VERSION : 1.4
// Der FC 53 kann fuer Motoren mit Umrichter, 2 Drehzahlen bzw 2 Punkteverstellung 
// verwendet werden.
// 
// Wird der Baustein mit Umrichter betrieben, so ist das Netzschuetz fuer den 
// Umrichter ans Netz verwendet.
// 
// Wir der Baustein ohne Umrichter betrieben, so ist das Netzschuetz fuer die  
// kleine Drehzahl verwendet.
// 
// Info: Stoerung Laufzeit Speisepumpe. Die eingestellte Zeit in der die 
// Speisepumpe den Pumpenvordruck aufbauen muss ist abgelaufen.
   VAR_INPUT
      IN_ControlVoltage : Bool;   // Delay switch on frequency unit after emergency stop (protection)
      IN_OperationMode_Valid : Bool;   // A valid operation mode (manual or automatic) is selected
      IN_OPerationMode_Active : Bool;   // Opearation mode is selected and hydraulic is active
      IN_Min_PrePressure : Bool;   // Inputsignal pressurelevel of pre pressure pump reached
      IN_Max_PressureComponent : Bool;   // Inputsignal maximum component pressure after pump exceeded
      IN_MotorprotectionPump : Bool;   // Inputsignal error power supply or motor protection of component pump
      IN_With_FU_Pump : Bool;   // Select control of component pump by frequeny unit
      IN_FLT_FU_Pump : Bool;   // Inputsignal fault of frequeny unit component pump
      IN_MaxLevelTray : Bool;   // Input fault max. filling level tray
      IN_Shot_Start : Bool;   // Foaming is active
      IN_MinPressure : Bool;   // Inputsignal fault min pressure of component pump
      IN_PreAlarmBearing : Bool;
      IN_AlarmBearing : Bool;
      IN_Reset_fault_Fkt : Bool;   // Quit faults inside the function block
      IN_ReleaseExternal : Bool;   // External Signal release of pump-/ frequncy unit
      IN_FaultGroup_1 : Bool;   // Fault message of level 1 is active and was not acknowledged
      IN_SOverSOffSWU_running : Bool;   // Switchover- Switchoff- time switch over unit still running
      IN_High_speed : Bool;   // High speed running
      IN_2point_Adjustment : Bool;   // 2 point adjustment is activ
      IN_Cycle_running : Bool;   // Foaming cycle was started and is active
      IN_Recirc_reduced : Bool;   // Reduced recirculation is selected and active
      IN_Recirc_lowpressure : Bool;   // Lowpressure recirculation is selected and active
      IN_Recirc_highpressure : Bool;   // Highpressure recirculation is selected and active
      IN_Recirc_pausetime : Bool;   // Pausetime during interval function active
      IN_UsedForShot : Bool;   // This component will be used for the next part shot
      IN_Delay_Restart : S5Time;   // Time value restart lock of component pump
      IN_Timer_Restart : Timer;   // Timer restart lock of component pump
      IN_RunDownTime_FeedPump : S5Time;   // Time value run down time feed pump
      IN_Timer_ControlFeedPump : Timer;   // Timer of pressure build up control feed pump
      IN_TimerOffFeedPump : Timer;   // Timer to delay switch off from feeding pump
      IN_Timer_Delay_EnClosedL : Timer;   // Timer delay release flow controller
      IN_TimerInterval : Timer;   // Timer for interval times
   END_VAR
   VAR_OUTPUT
      OUT_2_Point_Adjust : Bool;   // Output 2 point adjustment of pump
      OUT_Dosing_active : Bool;   // Signal dosing of component to ProCan-modul
      OUT_Enableclosedloop : Bool;   // Signal of Flow Index "enableclosedloop" to ProCan-modul
      OUT_Pump_MainsContactor : Bool;   // Output mainscontactor pump/frequency unit; or low speed contactor
      OUT_Release_FU : Bool;   // Output release frequency unit; or high speed contactor
   END_VAR
   VAR_IN_OUT
      IO_QPB_Pumpe : Bool;   // Toggelsignal of quick pressure build up to ProCan modul
      IO_Status : ANY;   // Storage of state component pump - state of program block
      IO_Fault : ANY;
      IO_Config : ANY;
      IO_NewFault : Bool;
      IO_FaultLevel_1 : Bool;
      IO_FaultLevel_2 : Bool;
      IO_FaultLevel_3 : Bool;
   END_VAR
   VAR_TEMP
      Temp_IO_Status : "UDT053_Pump";
      ERROR_CODE : Int;   // Error state of systemfunction "BLKMOV" Blockmove
      AnyPointer1 : ANY;   // Pointer to copy the array "IO_Status" and "Temp_IO_Status"
      AnyPointer2 : ANY;   // Pointer to copy the array "IO_Status" and "Temp_IO_Status"
      AnyPointer3 : ANY;   // Pointer to copy the array "IO_Config"
      ReleaseFentingPump : Bool;   // Flag of release fenting pump
      Feedpump_wo_postrun : Bool;   // Flag activation feed pump without component pump post run
      Temp_IO_Fault : "UDT1853_FLT_MeteringPump";
      Temp_IO_Config : "UDT753_MeteringPump";
      ComponentOFF : Bool;   // Component is switched off or on pause time interval
   END_VAR
BEGIN

REGION Network 1: Saved data integration
   // Änderungen:
   // -------------------------------------------------------------------------------
   // Da nach einem sofortigem Widereinschalten der Pumpen nach einer Störung 
   // "STG_Max_Druck" kann es zu einem beschädigen der Pumpen kommen. 
   // Hier wird hier nun über den Weg der Entlüftungspumpe eine Einschaltverzögerung 
   // vorgenommen.
   // 
   // v.d.Geest     20.09.2005
   // -------------------------------------------------------------------------------
   // Auch wenn die Pumpe nicht mit Speisepumpe betrieben wurde wird das Bit 
   // "#Temp_IO_Status.Anforderung_Speisepumpe" gesetzt. 
   // Dieses Signal wurde direkt mit dem Eingang "#IN_Mit_Speisepumpe" verknüpft.
   // 
   // v.d.Geest     16.07.2005
   // -------------------------------------------------------------------------------
   // Der Ausgang "OUT_hohe_Drehzahl" kann entfallen wenn dieser mit dem Ausgang 
   // "#OUT_Freigabe_an_FU_Pumpe" zusammengelegt wird.
   // Bei einem Pumpenstrang ohne Umrichter wäre dieses nun der Ausgang für die hohe 
   // Drehzahl der Pumpen.
   // 
   // Escher        25.11.2004
   // -------------------------------------------------------------------------------
   // Das Signal "Dosieren_an_PUC" war von der Reglerfreigabe an den 
   // Frequenzumrichter abhängig. Die PUC benötigt dieses Signal aber im Schäumzyklus 
   // auch bei ungeregelten Maschinen. (Änderungen im Netzwerk 7)
   // 
   // Strauß        02.08.2004
   // -------------------------------------------------------------------------------
   // Bei einer Verwendung der Komponentenpumpe mit Speisepumpe trat beim ausschalten 
   // der Betriebsart im Kreislauf die Störung "STG_SpP_Laufzeit" auf.
   // Dieses war der Fall wenn die Nachlaufzeit größer eingegeben war als die 
   // Überwachungszeit des Vordrucks.
   // Dieses wurde unterbunden indem die Speisepumpe bei nicht aktiver Betriebsart 
   // nicht mehr angesteuert wird. 
   // Änderungen im Netzwerk 5 durch einfügen von "#IN_Betriebsart_Aktiv" bei der 
   // Zuweisung der "#Temp_IO_Status.Anforderung_Speisepumpe".
   // 
   // v.d.Geest     09.09.2003
   // -------------------------------------------------------------------------------
   // Wenn die Komponentenpumpe ohne Umrichter betrieben wird ist es nicht nötig das 
   // die Anlaufverzögerung nach Steuerspannung Aus abläuft.
   // Deshalb wird das Bit "FRG_UR_wieder_ans_Netz" auch gesetzt, wenn kein Umrichter 
   // verwendet wird. Hierdurch brauch auch die Freigabe für den Zyklus nicht 
   // verändert werden.
   // 
   // v.d.Geest     15.04.2003
   // -------------------------------------------------------------------------------
   // Wenn mehrere Komponentenpumpen mit Speise- oder Entlüftungspumpen betrieben 
   // werden konnte ein unterschiedliches Anlaufen der Komponentenpumpen nur 
   // "außerhalb" des Bausteins unterbunden werden.
   // Hierfür wurde der neue Übergabeparameter "IN_Freigabe_extern" eingebunden. Also 
   // bitte bei einspielen des Bausteins auf die Änderung bim FB achten.
   // 
   // v.d.Geest     11.04.2003
   // -------------------------------------------------------------------------------
   // Um bei größeren Komponentenpumpen auch beim Ausschalten des Kreislaufes oder 
   // nach dem Zyklus ein nichtabreißen des Komponentenstromes zu gewährleisten muß 
   // hier die Speisepumpe, falls vorhanden, nachlaufen.
   // Diese Nachlaufzeit wird von außen vorgegeben sollte aber "fest" bleiben.
   // 
   // Jäger         01.04.2003
   // -------------------------------------------------------------------------------
   // Bei unterschreiten des Min. Füllstandes während des Zyklusses wurde die 
   // Ansteuerung der Materialpumpen abgebrochen.
   // Nur noch ein Abbruch wenn der Zyklus nicht mehr läuft
   // 
   // v.d.Geest     25.02.2003
   // -------------------------------------------------------------------------------
   // Die Störung des Vordruckes wird unabhängig von der Anforderung ausgewertet.
   // Hierdurch wird ein kurzes Anlaufen der Materialpumpnen bei nicht vorhandenen 
   // Vordruck unterbunden.
   // 
   // Lindner       27.01.2003
   // -------------------------------------------------------------------------------
         LAR1;
         L;
         LAR2;
   //
         L     W[AR2, P#0.0];  // Bytes
         T     W[AR1, P#0.0];
         L     W[AR2, P#2.0];  //Amount of bytes
         T     W[AR1, P#2.0];
         L     W[AR2, P#4.0];  //Block no,
         T     W[AR1, P#4.0];
         L     D[AR2, P#6.0];  //Startadress of datas
         T     D[AR1, P#6.0];
   //
         CALL  BLKMOV
         ( SRCBLK  := #AnyPointer1,
           RET_VAL := #ERROR_CODE,
           DSTBLK  := #Temp_IO_Status
         );
   //
         LAR1;
         L;
         LAR2;
   //
         L     W[AR2, P#0.0];  // Bytes
         T     W[AR1, P#0.0];
         L     W[AR2, P#2.0];  //Amount of bytes
         T     W[AR1, P#2.0];
         L     W[AR2, P#4.0];  //Block no,
         T     W[AR1, P#4.0];
         L     D[AR2, P#6.0];  //Startadress of datas
         T     D[AR1, P#6.0];
   //
         CALL  BLKMOV
         ( SRCBLK  := #AnyPointer2,
           RET_VAL := #ERROR_CODE,
           DSTBLK  := #Temp_IO_Fault
         );
   //
   //
         LAR1;
         L;
         LAR2;
   //
         L     W[AR2, P#0.0];  // Bytes
         T     W[AR1, P#0.0];
         L     W[AR2, P#2.0];  //Amount of bytes
         T     W[AR1, P#2.0];
         L     W[AR2, P#4.0];  //Block no,
         T     W[AR1, P#4.0];
         L     D[AR2, P#6.0];  //Startadress of datas
         T     D[AR1, P#6.0];
   //
         CALL  BLKMOV
         ( SRCBLK  := #AnyPointer3,
           RET_VAL := #ERROR_CODE,
           DSTBLK  := #Temp_IO_Config
         );
END_REGION

REGION Network 2: Handle interval mode
   // Messages
         A     #Temp_IO_Config.PumpDeselectedInterval;
         FP    #Temp_IO_Status.Mes_PumpDeselectedInt;
         R     #Temp_IO_Config.PumpDeselected;
         A     #Temp_IO_Config.PumpDeselected;
         FP    #Temp_IO_Status.Mes_PumpDeselected;
         R     #Temp_IO_Config.PumpDeselectedInterval;

         A     #Temp_IO_Status.Mes_PumpDeselectedInt;
         =     #Temp_IO_Fault.Mes_PumpDeselectedInt;
         A     #Temp_IO_Status.Mes_PumpDeselected;
         =     #Temp_IO_Fault.Mes_PumpDeselected;

         AN    #Temp_IO_Config.PumpDeselectedInterval;
         R     #Temp_IO_Status.IntervalPause;

   // Interval times
         A     #Temp_IO_Config.PumpDeselectedInterval;
         FP    #Temp_IO_Status.HF_FPPumpDeselectedInt;
         JCN   int;
         R     #Temp_IO_Status.IntervalPause;
         CLR;
         L     S5T#0MS;
         SP    #IN_TimerInterval;
         JU    eint;

   int:  AN    #Temp_IO_Config.PumpDeselectedInterval;
         JC    eint;

   // Change run time <-> pause time
         AN    #IN_TimerInterval;
         JCN   eint;

   // Select the correct time
         L     #Temp_IO_Config.RunTimePumpInterval;
         A     #Temp_IO_Status.IntervalPause;
         JC    time;
         L     #Temp_IO_Config.PauseTimePumpInterval;

   // Start timer
   time: CLR;
         SE    #IN_TimerInterval;
         SET;
         SE    #IN_TimerInterval;
         AN    #Temp_IO_Status.IntervalPause;
         =     #Temp_IO_Status.IntervalPause;
   eint: NOP   0;
   // switch off if necessary
         O     #Temp_IO_Config.PumpDeselected;
         O     #Temp_IO_Status.IntervalPause;
         =     #ComponentOFF;
END_REGION

REGION Network 3: Switch on delay of frequency unit
   // Bei Betrieb mit Umrichter wird der Umrichter mit einer Wiedereinschaltsperre 
   // von 30 Sek. geschützt. Nach Steuerspannung AUS wird der Umrichter 30 Sek. lang 
   // vom Netz getrennt auch wenn die Steuerspannung sofort wieder eingeschaltet 
   // wird.
   //--------- Frequency unit back to power supply ---------------
   //      O     #Temp_IO_Status.FLT_Max_pressure    // Bitte testen 25.6.08 HK
         AN    #IN_ControlVoltage;
         AN    #ComponentOFF;
         O     #ComponentOFF;
         FP    #Temp_IO_Status.Rampe_Voltage_Off;
         R     #Temp_IO_Status.Release_Startup_FC;
         R     #IN_Timer_Restart;
         R     #Temp_IO_Status.Start_Startupdelay;
   //
         A     #Temp_IO_Status.Release_Startup_FC;
         JC    Run;
   //
         A     #Temp_IO_Status.Start_Startupdelay;
         AN    #Temp_IO_Status.Release_Startup_FC;
         L     S5T#10S;
         SD    #IN_Timer_Restart;
   //
         SET;
         S     #Temp_IO_Status.Start_Startupdelay;
   //
         O     #IN_Timer_Restart;
         ON    #IN_With_FU_Pump;
         S     #Temp_IO_Status.Release_Startup_FC;
         R     #IN_Timer_Restart;
         R     #Temp_IO_Status.Start_Startupdelay;
   //
   Run:  NOP   0;
END_REGION

REGION Network 4: Fault handling
   //--------- Störung Reset --------------------------
         A     #IN_Reset_fault_Fkt;
         R     #Temp_IO_Fault.FLT_Prepressure;
         R     #Temp_IO_Fault.FLT_Motorprotection;
         R     #Temp_IO_Fault.FLT_Max_pressure;
         R     #Temp_IO_Fault.FLT_SpP_Runtime;
         R     #Temp_IO_Fault.FLT_F_converter;
         R     #Temp_IO_Fault.FLT_Min_Pressure;
         R     #Temp_IO_Fault.FLT_DeselectedCompReqest;
         R     #Temp_IO_Fault.FLT_MaxLTripTray;
         R     #Temp_IO_Fault.FLT_PreAlarmBearing;
         R     #Temp_IO_Fault.FLT_AlarmBearing;
   //--------- Störung Pumpenvordruck -----------------
         A     #Temp_IO_Status.Netrelais;
         AN    #IN_Min_PrePressure;
         AN    #IN_With_FU_Pump;
         O;
         A     #IN_With_FU_Pump;
         A     #Temp_IO_Status.Controllrelease_to_FC;
         AN    #IN_Min_PrePressure;
         O;
         AN    #Temp_IO_Config.WithFeedPump;
         AN    #IN_Min_PrePressure;
         AN    #ComponentOFF;
         AN    #Temp_IO_Fault.FLT_Prepressure;
         S     #Temp_IO_Fault.FLT_Prepressure;
         S     #IO_NewFault;
   //--------- Störung Laufzeit Speisepumpe -----------
         A     #Temp_IO_Status.Selection_Feedingpump;
         A     #Temp_IO_Config.WithFeedPump;
         AN    #IN_Min_PrePressure;
         L     #Temp_IO_Config.DelayPressureFeedP;
         SD    #IN_Timer_ControlFeedPump;
   //
         A     #IN_Timer_ControlFeedPump;
         AN    #Temp_IO_Fault.FLT_SpP_Runtime;
         S     #Temp_IO_Fault.FLT_SpP_Runtime;
         S     #IO_NewFault;
   //--------- Störung Motorschutz --------------------
         A     #IN_MotorprotectionPump;
         AN    #ComponentOFF;
         AN    #Temp_IO_Fault.FLT_Motorprotection;
         S     #Temp_IO_Fault.FLT_Motorprotection;
         S     #IO_NewFault;
   //--------- Störung max. Druck  --------------------
         AN    #IN_Max_PressureComponent;
         AN    #ComponentOFF;
         AN    #Temp_IO_Fault.FLT_Max_pressure;
         S     #Temp_IO_Fault.FLT_Max_pressure;
         S     #IO_NewFault;
   //--------- Fault deselected component requested for shot  ---
         O     #Temp_IO_Config.PumpDeselectedInterval;
         O     #Temp_IO_Config.PumpDeselected;
         A     #IN_UsedForShot;
         AN    #Temp_IO_Fault.FLT_DeselectedCompReqest;
         S     #Temp_IO_Fault.FLT_DeselectedCompReqest;
         S     #IO_NewFault;
   //--------- Störung Umrichter  ---------------------
         ON    #IN_With_FU_Pump;
         ON    #Temp_IO_Status.Release_Startup_FC;
         O     #ComponentOFF;
         JC    K_UR;
         A     #Temp_IO_Status.Netrelais;
         L     S5T#15S;
         SD    #IN_Timer_Restart;
         A     #IN_Timer_Restart;
         AN    #IN_FLT_FU_Pump;
         AN    #Temp_IO_Fault.FLT_F_converter;
         S     #Temp_IO_Fault.FLT_F_converter;
         S     #IO_NewFault;

   //-----
         AN    #IN_MaxLevelTray;
         AN    #Temp_IO_Fault.FLT_MaxLTripTray;
         S     #Temp_IO_Fault.FLT_MaxLTripTray;
         S     #IO_NewFault;

   K_UR: NOP   0;
   //--------- Min pressure at     -------------------
   //---------  shot start         -------------------
         A     #IN_Shot_Start;
         AN    #IN_MinPressure;
         A     #IN_UsedForShot;
         AN    #Temp_IO_Fault.FLT_Min_Pressure;
         S     #Temp_IO_Fault.FLT_Min_Pressure;
         S     #IO_NewFault;

         A     #IN_PreAlarmBearing;
         AN    #Temp_IO_Fault.FLT_PreAlarmBearing;
         S     #Temp_IO_Fault.FLT_PreAlarmBearing;
         S     #IO_NewFault;

         A     #IN_AlarmBearing;
         AN    #Temp_IO_Fault.FLT_AlarmBearing;
         S     #Temp_IO_Fault.FLT_AlarmBearing;
         S     #IO_NewFault;

         A     #Temp_IO_Status.Start_Startupdelay;
         =     #Temp_IO_Fault.Mes_StartUpDelayFU;
END_REGION

REGION Network 5: Error handling fault groups
         O     #Temp_IO_Fault.FLT_Prepressure;
         O     #Temp_IO_Fault.FLT_Motorprotection;
         O     #Temp_IO_Fault.FLT_Max_pressure;
         O     #Temp_IO_Fault.FLT_F_converter;
         O     #Temp_IO_Fault.FLT_SpP_Runtime;
         O     #Temp_IO_Fault.FLT_Min_Pressure;
         O     #Temp_IO_Fault.FLT_DeselectedCompReqest;
         O     #Temp_IO_Fault.FLT_AlarmBearing;
         O     #Temp_IO_Fault.FLT_MaxLTripTray;
         S     #IO_FaultLevel_1;

   //      O     XXXXXXXX
   //      S     #IO_FaultLevel_2

         O     #Temp_IO_Fault.FLT_PreAlarmBearing;
         S     #IO_FaultLevel_3;
   //
         O     #Temp_IO_Fault.FLT_Prepressure;
         O     #Temp_IO_Fault.FLT_Motorprotection;
         O     #Temp_IO_Fault.FLT_Max_pressure;
         O     #Temp_IO_Fault.FLT_F_converter;
         O     #Temp_IO_Fault.FLT_SpP_Runtime;
         O     #Temp_IO_Fault.FLT_Min_Pressure;
         O     #Temp_IO_Fault.FLT_DeselectedCompReqest;
         O     #Temp_IO_Fault.FLT_AlarmBearing;
         O     #Temp_IO_Fault.FLT_PreAlarmBearing;
         O     #Temp_IO_Fault.FLT_MotorFan;
         O     #Temp_IO_Fault.FLT_MaxLTripTray;
         =     #Temp_IO_Status.FLT_Exist;
END_REGION

REGION Network 6: Venting pump
   //       ON    #Temp_IO_Status.STG_Min_Level
   //       O     #IN_Cycle_running
   //     U     #IN_Mit_Entlueftungspumpe
   //       U     #IN_OperationMode_Valid
   //       UN    #Temp_IO_Fault.FLT_Prepressure
   //       =     #Freigabe_Enlt_Pumpe
   //
   //      U     #Temp_IO_Status.Ventingtime_finished
   //      SPB   P_ok
   //
   //      U     #Freigabe_Enlt_Pumpe
   //      L     S5T#10S
   //      SE    #IN_Timer_Universal
   //-------------------------------------------------
   //       O     #IN_Timer_Universal
   //       ON    #IN_Mit_Entlueftungspumpe
   //       S     #Temp_IO_Status.Ventingtime_finished
   //-------------------------------------------------
   //      SPBN  P_ok
   //
   //       CLR
   //       SI    #IN_Timer_Universal
   //
   // P_ok: NOP 0
   //-------------------------------------------------
   //       U     #Temp_IO_Status.STG_Min_Level
   //       UN    #IN_Cycle_running
   //       ON    #IN_ControlVoltage
   //       O     #Temp_IO_Fault.FLT_Prepressure
   //       R     #Temp_IO_Status.Ventingtime_finished
   //-------------------------------------------------
   //      ON    #Temp_IO_Status.Ventingtime_finished
   //       O     #Temp_IO_Status.Allg_Pumpenanforderung
   //       U     #Freigabe_Enlt_Pumpe
   //       UN    #Temp_IO_Status.STG_Motorsch_Entl_Pumpe
   //       =     #Temp_IO_Status.Netzschuetz_Entl_Pumpe
END_REGION

REGION Network 7: Pump
         O     #IN_Recirc_reduced;
         O     #IN_Recirc_lowpressure;
         A(;
         ON    #IN_Recirc_pausetime;
         O     #IN_Cycle_running;
         );
         O     #IN_Recirc_highpressure;
         O     #IN_Cycle_running;
         A     #IN_OPerationMode_Active;
         AN    #IN_FaultGroup_1;
         AN    #Temp_IO_Fault.FLT_Prepressure;
         AN    #Temp_IO_Fault.FLT_Motorprotection;
         AN    #Temp_IO_Fault.FLT_Max_pressure;
         AN    #Temp_IO_Fault.FLT_SpP_Runtime;
         AN    #Temp_IO_Fault.FLT_F_converter;
   //      U     #Temp_IO_Status.Ventingtime_finished
         A     #IN_ControlVoltage;
         AN    #ComponentOFF;
         =     #Feedpump_wo_postrun;
         A     #Feedpump_wo_postrun;
         L     #IN_RunDownTime_FeedPump;
         SF    #IN_TimerOffFeedPump;
   //
         A     #IN_TimerOffFeedPump;
         A     #Temp_IO_Config.WithFeedPump;
         A     #IN_OPerationMode_Active;
         =     #Temp_IO_Status.Selection_Feedingpump;
   //-------------------------------------------------
         ON    #Temp_IO_Status.Release_Startup_FC;
         O     #IN_With_FU_Pump;
         JC    Allg;
         AN    #IN_With_FU_Pump;
         A     #Temp_IO_Status.High_rpm;
         AN    #IN_High_speed;
         L     #IN_Delay_Restart;
         SE    #IN_Timer_Restart;
   //-------------------------------------------------
   Allg: AN    #IN_With_FU_Pump;
         A     #Feedpump_wo_postrun;
         A     #IN_Min_PrePressure;
         AN    #IN_Timer_Restart;
         O;
         A     #IN_With_FU_Pump;
         A     #Feedpump_wo_postrun;
         A     #IN_Min_PrePressure;
         =     #Temp_IO_Status.Main_Pumpselection;
   //------ Umrichter ans Netz bzw. kleine Drehzahl --
         A     #IN_ReleaseExternal;
         A     #Temp_IO_Status.Main_Pumpselection;
         AN    #IN_With_FU_Pump;
         O;
         A     #IN_With_FU_Pump;
         A     #IN_ControlVoltage;
         AN    #ComponentOFF;
         A     #Temp_IO_Status.Release_Startup_FC;
         =     #Temp_IO_Status.Netrelais;
   //-------------------------------------------------
         O     #IN_Recirc_reduced;
         O     #IN_Recirc_lowpressure;
         A(;
         ON    #IN_Recirc_pausetime;
         O     #IN_Cycle_running;
         );
         O     #IN_Recirc_highpressure;
         O     #IN_Cycle_running;
         A     #IN_ReleaseExternal;
         A     #Temp_IO_Status.Main_Pumpselection;
         AN    #Temp_IO_Fault.FLT_Prepressure;
         AN    #Temp_IO_Fault.FLT_Motorprotection;
         AN    #Temp_IO_Fault.FLT_Max_pressure;
         AN    #Temp_IO_Fault.FLT_SpP_Runtime;
         AN    #Temp_IO_Fault.FLT_F_converter;
         A     #IN_FLT_FU_Pump;
         =     #Temp_IO_Status.Controllrelease_to_FC;
END_REGION

REGION Network 8: High speed and 2 point adjustment if drive without FU
         A     #Temp_IO_Status.Netrelais;
         A     #IN_High_speed;
         =     #Temp_IO_Status.High_rpm;
   //-------------------------------------------------
         A     #Feedpump_wo_postrun;
         A     #IN_2point_Adjustment;
         =     #Temp_IO_Status.Valve_2_point_selection;
END_REGION

REGION Network 9: Release of controller to modul of machine
         A     #IN_ReleaseExternal;
         A     #Temp_IO_Status.Main_Pumpselection;
         AN    #IN_With_FU_Pump;
         O     #Temp_IO_Status.Controllrelease_to_FC;
         =     #Temp_IO_Status.Metering_to_PUC;
   //
         A     #Temp_IO_Status.Controllrelease_to_FC;
         L     S5T#300MS;
         SD    #IN_Timer_Delay_EnClosedL;

         A     #IN_Timer_Delay_EnClosedL;
         =     #Temp_IO_Status.Enableclosedloop;
END_REGION

REGION Network 10: Quick pressure build up
   // Nur notwendig fuer "Schnellen Druckaufbau" mit Modul !!!
         O     #IN_Cycle_running;
         O     #IN_Recirc_highpressure;
         A     #IN_With_FU_Pump;
         AN    #IN_SOverSOffSWU_running;
         A     #Temp_IO_Status.Enableclosedloop;
         A(;
         O     #IN_UsedForShot;
         ON    #IN_Cycle_running;
         );
         FP    #Temp_IO_Status.Puls_SDA;
         JCN   SDA;
         AN    #IO_QPB_Pumpe;
         =     #IO_QPB_Pumpe;
   SDA:  NOP   0;
END_REGION

REGION Network 11: Allocation of outputs
         A     #Temp_IO_Status.Netrelais;
         =     #OUT_Pump_MainsContactor;
   //-------------------------------------------------
         A     #Temp_IO_Status.Valve_2_point_selection;
         =     #OUT_2_Point_Adjust;
   //-------------------------------------------------
         A     #Temp_IO_Status.Controllrelease_to_FC;
         A     #IN_With_FU_Pump;
         O;
         A     #Temp_IO_Status.High_rpm;
         AN    #IN_With_FU_Pump;
         =     #OUT_Release_FU;
   //-------------------------------------------------
         A     #Temp_IO_Status.Metering_to_PUC;
         =     #OUT_Dosing_active;
   //-------------------------------------------------
         A     #IN_With_FU_Pump;
         A     #Temp_IO_Status.Enableclosedloop;
         =     #OUT_Enableclosedloop;
   //-------------------------------------------------
END_REGION

REGION Network 12: Function is active
         SET;
         =     #Temp_IO_Status.Block_is_active;
END_REGION

REGION Network 13: Save data
         CALL  BLKMOV
         ( SRCBLK  := #Temp_IO_Status,
           RET_VAL := #ERROR_CODE,
           DSTBLK  := #AnyPointer1
         );
   //
         CALL  BLKMOV
         ( SRCBLK  := #Temp_IO_Fault,
           RET_VAL := #ERROR_CODE,
           DSTBLK  := #AnyPointer2
         );
   //
         CALL  BLKMOV
         ( SRCBLK  := #Temp_IO_Config,
           RET_VAL := #ERROR_CODE,
           DSTBLK  := #AnyPointer3
         );
END_REGION
END_FUNCTION

FUNCTION "FC054_FaultsMetering" : Void   // FC54, STL
TITLE = Faults ProCan flowstate
{ S7_Optimized_Access := 'FALSE' }
NAME : Fault
VERSION : 0.1
   VAR_INPUT
      IN_ProCanFlow_State : Struct
         Flowstopped : Bool;   // piston has stopped
         FlowQPB : Bool;   // Flow quick pressure build up is active
         ControlOnUpperLimit : Bool;   // flow control loop operates on it upper limits
         ControlOnLowerLimit : Bool;   // flow control loop operates on its lower limits
         FlowtoleranceL : Bool;   // tolerance: flow is too low
         FlowtoleranceH : Bool;   // tolerance: flow is too high
      END_STRUCT;
      IN_Reset_Fault : Bool;
   END_VAR
   VAR_IN_OUT
      IO_Any_Flow_Fault : ANY;
      IO_HF_FLT_QPB : Bool;
      IO_FaultLevel1 : Bool;
      IO_FaultLevel2 : Bool;
      IO_FaultLevel3 : Bool;
      IO_NewFault : Bool;
   END_VAR
   VAR_TEMP
      Temp_Any_Flow_Fault : ANY;
      Temp_Flow_Fault : "UDT1853_FLT_MeteringPump";
      ERROR_CODE : Int;
      Temp_FLT_Tolerance_high : Bool;
      Temp_FLT_Tolerance_low : Bool;
      Temp_FLT_FlowContrAtLim : Bool;
      Temp_Flt_FlowSDAtimeOut : Bool;
   END_VAR
BEGIN

REGION Network 1: Get temporary variables flow fault
         L;
         LAR1;
         LAR2;
   //
         L     W[AR1, P#0.0];  // Bytes
         T     W[AR2, P#0.0];
         L     W[AR1, P#2.0];  // Amount of bytes
         T     W[AR2, P#2.0];
         L     W[AR1, P#4.0];  // Block no,
         T     W[AR2, P#4.0];
         L     D[AR1, P#6.0];  // Startadress of data
         T     D[AR2, P#6.0];
   //
         CALL  BLKMOV
         ( SRCBLK  := #Temp_Any_Flow_Fault,
           RET_VAL := #ERROR_CODE,
           DSTBLK  := #Temp_Flow_Fault
         );
END_REGION

REGION Network 2: Reset faults flow
         AN    #IN_Reset_Fault;
         JC    nw3e;

         CLR;
         =     #Temp_Flow_Fault.FLT_Tolerance_high;
         =     #Temp_Flow_Fault.FLT_Tolerance_low;
         =     #Temp_Flow_Fault.FLT_FlowControlAtLimit;
         =     #Temp_Flow_Fault.FLT_FlowControlAtLOWLimit;
         =     #Temp_Flow_Fault.FLT_FlowSDATimeOut;

   nw3e: NOP   0;
END_REGION

REGION Network 3: Fault flow state of ProCan module
   //      L     #IN_ProCanFlow_State
   //      L     16
   //      UW
   //      L     0
   //      <>D
   //      FP    #IO_HF_FLT_QPB
   //      =     #Temp_Flt_FlowSDAtimeOut

   //      U     #Temp_Flt_FlowSDAtimeOut
   //      UN    #Temp_Flow_Fault.FLT_FlowSDATimeOut
   //      S     #Temp_Flow_Fault.FLT_FlowSDATimeOut
   //      S     #IO_NewFault

         A     #IN_ProCanFlow_State.ControlOnUpperLimit;
         AN    #Temp_Flow_Fault.FLT_FlowControlAtLimit;
         S     #Temp_Flow_Fault.FLT_FlowControlAtLimit;
         S     #IO_NewFault;

         A     #IN_ProCanFlow_State.ControlOnLowerLimit;
         AN    #Temp_Flow_Fault.FLT_FlowControlAtLOWLimit;
         S     #Temp_Flow_Fault.FLT_FlowControlAtLOWLimit;
         S     #IO_NewFault;
END_REGION

REGION Network 4: Fault levels
   //    O     xxxxxxxxx
   //    =     #IO_FaultLevel1

         O     #Temp_Flow_Fault.FLT_Tolerance_high;
         O     #Temp_Flow_Fault.FLT_Tolerance_low;
         O     #Temp_Flow_Fault.FLT_FlowControlAtLimit;
         O     #Temp_Flow_Fault.FLT_FlowControlAtLOWLimit;
         O     #Temp_Flow_Fault.FLT_FlowSDATimeOut;
         S     #IO_FaultLevel3;
END_REGION

REGION Network 5: Write back faults
         CALL  BLKMOV
         ( SRCBLK  := #Temp_Flow_Fault,
           RET_VAL := #ERROR_CODE,
           DSTBLK  := #Temp_Any_Flow_Fault
         );
END_REGION
END_FUNCTION

FUNCTION "FC055_PumpVentilation" : Void   // FC55, STL
TITLE = Function for organize pump Ventilation
{ S7_Optimized_Access := 'FALSE' }
VERSION : 0.1
   VAR_INPUT
      IN_Reset_fault_Fkt : Bool;   // Quit faults inside the function block
      IN_Motorprotection : Bool;   // Inputsignal error power supply or motor protection
      IN_ComponentDeselected : Bool;   // Is the component deselected? -> Fault Group 2 -> Groupe 3
      In_Start : Bool;   // Start value for the ventilation
      IN_Time : S5Time;   // Time value delay switch off the ventilation
      IN_Timer : Timer;   // Timer for delay time to switch off the ventilation
   END_VAR
   VAR_OUTPUT
      OUT_MainContactor : Bool;   // Output maincontactor Ventilation
   END_VAR
   VAR_IN_OUT
      IO_FLT_MotorFan : Bool;
      IO_NewFault : Bool;
      IO_FaultLevel_2 : Bool;
      IO_FaultLevel_3 : Bool;
   END_VAR
BEGIN

REGION Network 1: Fault handling
   //--------- Reset fault ---------------------------
         A     #IN_Reset_fault_Fkt;
         R     #IO_FLT_MotorFan;
   //--------- Fault Motorprotection -----------------
         A     #IN_Motorprotection;
         AN    #IO_FLT_MotorFan;
         S     #IO_FLT_MotorFan;
         S     #IO_NewFault;
   //--------- If selected fault group 2 -------------
         A     #IO_FLT_MotorFan;
         AN    #IN_ComponentDeselected;
         S     #IO_FaultLevel_2;
   //--------- If deselected fault group 3 -----------
         A     #IO_FLT_MotorFan;
         A     #IN_ComponentDeselected;
         S     #IO_FaultLevel_3;
   //-------------------------------------------------
END_REGION

REGION Network 2: Start venting
   //-----
         A     #In_Start;
         AN    #IO_FLT_MotorFan;
         L     #IN_Time;
         SF    #IN_Timer;
         A     #IN_Timer;
         AN    #IO_FLT_MotorFan;
         =     #OUT_MainContactor;
   //-----
END_REGION
END_FUNCTION

FUNCTION "FC056_TemPulse2" : Void   // FC56, STL
TITLE = Temperature control pulse width
{ S7_Optimized_Access := 'FALSE' }
VERSION : 0.1
   VAR_INPUT
      Trig : Bool;
      In_Sollwert : Real;
      In_Istwert_Tank : Real;
      In_Istwert_Return : Real;
      In_Wichtung : Real;
      In_Regelstrecke : Real;
      In_MaxDelta_K : Real;
      In_MaxDelta_H : Real;
   END_VAR
   VAR_IN_OUT
      Pulsezeit : Real;
      Heating : Bool;
      Cooling : Bool;
   END_VAR
   VAR_TEMP
      Value1 : Real;
      Value2 : Real;
      Value3 : Real;
      Value4 : Real;
      Value5 : Real;
      Value6 : Real;
      Value7 : Real;
      MaxDelta : Real;
      Istwert_Tank : Real;
      Istwert_Return : Real;
      Sollwert : Real;
      Wichtung : Real;
      MaxDelta_K : Real;
      MaxDelta_H : Real;
      Regelstrecke : Real;
      Pulsezeit_real : Real;
   END_VAR
BEGIN

REGION Network 1: Berechnen nur wenn Timer abgelaufen
         AN    #Trig;
         BEC;
END_REGION

REGION Network 2: Werte wandeln von INT in REAL
         L     #In_Sollwert;
         T     #Sollwert;

         L     #In_Istwert_Tank;
         T     #Istwert_Tank;

         L     #In_Istwert_Return;
         T     #Istwert_Return;

         L     #In_Wichtung;
         T     #Wichtung;

         L     #In_Regelstrecke;
         T     #Regelstrecke;

         L     #In_MaxDelta_K;
         T     #MaxDelta_K;

         L     #In_MaxDelta_H;
         T     #MaxDelta_H;
END_REGION

REGION Network 3: Mittelwert bilden
         L     #Istwert_Tank;
         L     #Wichtung;
         *R;
         T     #Value1;

         L     100.0;
         L     #Wichtung;
         -R;
         L     #Istwert_Return;
         *R;
         T     #Value2;

         L     #Value1;
         L     #Value2;
         +R;
         L     100.0;
         /R;
         T     #Value3;  // Mittelwert
END_REGION

REGION Network 4
   // Ist dieser Wert negativ, dann mit MaxDelta_H arbeiten
         L     #Value3;
         L     #Sollwert;
         -R;
         T     #Value4;  // Differenz Mittelist - Sollwert

         L     #MaxDelta_K;  // Wert für Kühlen
         T     #MaxDelta;

         L     #Value4;
         L     0;
         <R;
         JCN   Limi;
         L     #MaxDelta_H;  // Für Heizen diesen Wert nehmen
         T     #MaxDelta;
END_REGION

REGION Network 5
   // Differenz auf MaxWert limitieren
   Limi: L     #Value4;
         L     #MaxDelta;
         >R;
         JCN   kMax;
         T     #Value5;
         JU    calc;

   kMax: L     #Value4;
         T     #Value5;
END_REGION

REGION Network 6
   calc: NOP   0;

         L     100.0;
         L     #Value5;
         *R;
         L     #MaxDelta;
         /R;
         T     #Value6;
END_REGION

REGION Network 7: Pulsezeit: - >> HEIZEN / + >> KÜHLEN
         L     #Regelstrecke;
         L     100.0;
         /R;
         L     #Value6;
         *R;
         T     #Value7;

         L     #Value7;
         L     100.0;
         *R;
         T     #Pulsezeit_real;

   // Wenn noch nicht Positiv, dann machen !
         L     #Pulsezeit_real;
         L     0.0;
         <R;
         JCN   tak;
         L     #Pulsezeit_real;
         NEGR;
         JU    rnd;

   tak:  TAK;
   rnd:  NOP   0;
         L     10.0;
         *R;
         T     #Pulsezeit;  // Ausgabe int INT, aber gleich positiv!
END_REGION

REGION Network 8: Steuerbits ausgeben
         L     #Pulsezeit_real;
         L     0.0;
         >R;
         =     #Cooling;

         L     #Pulsezeit_real;
         L     0.0;
         <R;
         =     #Heating;
END_REGION
END_FUNCTION

FUNCTION "FC057_HPHeatexchanger" : Void   // FC57, STL
{ S7_Optimized_Access := 'FALSE' }
VERSION : 0.1
   VAR_TEMP
      DINT_dummy : Real;
      Imp_WT_Aus : Bool;
      Imp_WT_Ein : Bool;
      Temp_Cooling : Bool;
      Dummy : Bool;
      Temp_MoreDelta : Bool;
      Temp_HD_WT : Real;
      Temp_SetValueTemp : Real;
      Regelstrecke : Time;
      Zeit_abgelaufen : Time;
   END_VAR
BEGIN

REGION Network 1: There is no connection to the sensor (3)
   //---------------------------------------------
   //  Controller temperature Heatexchanger K1
   //---------------------------------------------
         AN    "DB753_MeteringPump".Pump[1].WithHPHeatExchanger;
         R     "DB823_Error_Metering".Temperature_HeatexchangerHP[1].Sensor_FLT_broken_wire;
         R     "DB823_Error_Metering".Temperature_HeatexchangerHP[1].Warning_limit_plus;
         R     "DB823_Error_Metering".Temperature_HeatexchangerHP[1].Warning_limit_minus;
         R     "DB823_Error_Metering".Temperature_HeatexchangerHP[1].Alarm_limit_plus;
         R     "DB823_Error_Metering".Temperature_HeatexchangerHP[1].Alarm_limit_minus;
         R     "DB613_Komponent_State".HeatexchangerHP[1].Fault_Exist;
         JC    EHD1;
   //-----
         CALL  "FC920_PV_Calc_Act_Value"
         ( IN_Act_Value_read := TRUE,
           IN_Act_Value_ext  := FALSE,
           IN_Ext_Value      := #DINT_dummy,
           IN_Read_Double    := FALSE,
           IN_FLT_Needful    := 1,
           IN_FLT_Reset      := "DB009_Faults".Faults_Reset_FKT_M1,
           IO_Any_ArrayPV    := "DB608_PV_Metering".HeatexchangerHP[1],
           IO_Fault_Sensor   := "DB823_Error_Metering".Temperature_HeatexchangerHP[1].Sensor_FLT_broken_wire,
           IO_New_Fault      := "DB009_Faults".Faultschanging_M1,
           IO_FLT_Level_3    := "DB009_Faults".Faults_FKT_Grp_3_M1
         );

   //---------------------------------------------
   //  Controller temperature Heatexchanger K1
   //---------------------------------------------
         L     "DB608_PV_Metering".HeatexchangerHP[1].PV_ActV.Value;
         L     10.0;
         /R;
         T     #Temp_HD_WT;
   //
         L     "DB608_PV_Metering".HeatexchangerHP[1].PV_SetV.Value;
         L     10.0;
         /R;
         T     #Temp_SetValueTemp;
   //
         CALL  "FC056_TemPulse2"
         ( Trig              := "Start_Controler1_HP_K1",
           In_Sollwert       := #Temp_SetValueTemp,
           In_Istwert_Tank   := #Temp_HD_WT,
           In_Istwert_Return := #Temp_HD_WT,
           In_Wichtung       := "DB751_auxiliaryDriveMetering".HeatexchangerHP[1].Weighting_Temp,
           In_Regelstrecke   := "DB751_auxiliaryDriveMetering".HeatexchangerHP[1].PLC_Control_Area,
           In_MaxDelta_K     := "DB751_auxiliaryDriveMetering".HeatexchangerHP[1].Max_Temp_Diff_Cooling,
           In_MaxDelta_H     := "DB751_auxiliaryDriveMetering".HeatexchangerHP[1].Max_Temp_Diff_Heating,
           Pulsezeit         := "DB613_Komponent_State".HeatexchangerHP[1].PulsTime,
           Heating           := #Dummy,
           Cooling           := #Temp_Cooling
         );
   //
   //Regelstrecke ms Format
         L     "DB751_auxiliaryDriveMetering".HeatexchangerHP[1].PLC_Control_Area;
         L     1000.0;
         *R;
         RND;
         T     #Regelstrecke;  // Zeitwert für Timer

   // Regelstreckentimer ständig starten

         AN    "Start_Controler1_HP_K1";
         =     "Start_Controler2_HP_K1";

         CALL  TON , "DB55_Temp_HD_WT_MK1_K1"
         ( IN := "Start_Controler2_HP_K1",
           PT := #Regelstrecke,
           Q  := "Start_Controler1_HP_K1",
           ET := #Zeit_abgelaufen
         );

   // Kühlen  EIN
         A     #Temp_Cooling;
         S     "DB613_Komponent_State".HeatexchangerHP[1].CoolingActive;

   // Kleine Einschatverzögerung
         L     #Temp_SetValueTemp;
         L     "DB751_auxiliaryDriveMetering".HeatexchangerHP[1].Offset_Cooling;
         +R;
         L     #Temp_HD_WT;
         >R;
         =     #Temp_MoreDelta;
   // Kühlen  AUS
         L     "DB613_Komponent_State".HeatexchangerHP[1].PulsTime;
         RND;
         L     #Zeit_abgelaufen;
         <D;
         AN(;
         L     "DB613_Komponent_State".HeatexchangerHP[1].PulsTime;
         RND;
         L     #Regelstrecke;
         >D;
         );
         ON    "DB613_Komponent_State".HeatexchangerHP[1].Switch_Temp_ON_OFF;
         ON    "DB619_State_MPart".Operationmode[1].valid;
         O     "DB823_Error_Metering".Temperature_HeatexchangerHP[1].Sensor_FLT_broken_wire;
         O     #Temp_MoreDelta;
         R     "DB613_Komponent_State".HeatexchangerHP[1].CoolingActive;

         A     "DB613_Komponent_State".HeatexchangerHP[1].CoolingActive;
         A     "DB619_State_MPart".Machine[1].Metering."01";

         =     "V_HP_Heater_Cooling_C1";  // "V_HExchang_Cooling_K1" // stromlos zu
         =     "V_HP_Heater_Bypass_C1";  // "V_HExchang_Bypass_K1" // stromlos offen

   //-----
   // Check limits temperature 1 Heatexchanger

         CALL  "FC916_PV_Limits"
         ( IN_Tolerance_Test     := "DB619_State_MPart".Operationmode[1].Controllvoltage,
           IN_Reset_Fault        := "DB009_Faults".Faults_Reset_FKT_M1,
           IO_Any_ArrayPV        := "DB608_PV_Metering".HeatexchangerHP[1],
           IO_Fault_Warn_upperL  := "DB823_Error_Metering".Temperature_HeatexchangerHP[1].Warning_limit_plus,
           IO_Fault_Warn_lowerL  := "DB823_Error_Metering".Temperature_HeatexchangerHP[1].Warning_limit_minus,
           IO_Fault_Alarm_upperL := "DB823_Error_Metering".Temperature_HeatexchangerHP[1].Alarm_limit_plus,
           IO_Fault_Alarm_lowerL := "DB823_Error_Metering".Temperature_HeatexchangerHP[1].Alarm_limit_minus,
           IO_New_Fault          := "DB009_Faults".Faultschanging_M1,
           IO_Fault_Level_1      := "DB009_Faults".Faults_FKT_Grp_1_M1,
           IO_Fault_Level_2      := "DB009_Faults".Faults_FKT_Grp_2_M1,
           IO_Fault_Level_3      := "DB009_Faults".Faults_FKT_Grp_3_M1
         );
   //-----
   // State of Switch
         L     0;
         A     "DB613_Komponent_State".HeatexchangerHP[1].CoolingActive;
         A     "DB619_State_MPart".Machine[1].Metering."01";
         A     "DB613_Komponent_State".HeatexchangerHP[1].Switch_Temp_ON_OFF;
         JCN   S1H1;
         L     1;
   S1H1: ON    "DB613_Komponent_State".HeatexchangerHP[1].CoolingActive;
         ON    "DB619_State_MPart".Machine[1].Metering."01";
         A     "DB613_Komponent_State".HeatexchangerHP[1].Switch_Temp_ON_OFF;
         JCN   S2H1;
         L     3;
   S2H1: A     "DB823_Error_Metering".Temperature_HeatexchangerHP[1].Sensor_FLT_broken_wire;
         A     "DB613_Komponent_State".HeatexchangerHP[1].Switch_Temp_ON_OFF;
         JCN   S3H1;
         L     2;
   S3H1: T     "DB613_Komponent_State".HeatexchangerHP[1].State_Temp;
   EHD1: NOP   0;

   // Fault exists
         O     "DB823_Error_Metering".Temperature_HeatexchangerHP[1].Sensor_FLT_broken_wire;
         O     "DB823_Error_Metering".Temperature_HeatexchangerHP[1].Warning_limit_plus;
         O     "DB823_Error_Metering".Temperature_HeatexchangerHP[1].Warning_limit_minus;
         O     "DB823_Error_Metering".Temperature_HeatexchangerHP[1].Alarm_limit_plus;
         O     "DB823_Error_Metering".Temperature_HeatexchangerHP[1].Alarm_limit_minus;
         =     "DB613_Komponent_State".HeatexchangerHP[1].Fault_Exist;
END_REGION

REGION Network 2: There is no connection to the sensor (3)
   //---------------------------------------------
   //  Controller temperature Heatexchanger K2
   //---------------------------------------------
         AN    "DB753_MeteringPump".Pump[2].WithHPHeatExchanger;
         R     "DB823_Error_Metering".Temperature_HeatexchangerHP[2].Sensor_FLT_broken_wire;
         R     "DB823_Error_Metering".Temperature_HeatexchangerHP[2].Warning_limit_plus;
         R     "DB823_Error_Metering".Temperature_HeatexchangerHP[2].Warning_limit_minus;
         R     "DB823_Error_Metering".Temperature_HeatexchangerHP[2].Alarm_limit_plus;
         R     "DB823_Error_Metering".Temperature_HeatexchangerHP[2].Alarm_limit_minus;
         R     "DB613_Komponent_State".HeatexchangerHP[2].Fault_Exist;
         JC    EHD2;
   //-----
         CALL  "FC920_PV_Calc_Act_Value"
         ( IN_Act_Value_read := TRUE,
           IN_Act_Value_ext  := FALSE,
           IN_Ext_Value      := #DINT_dummy,
           IN_Read_Double    := FALSE,
           IN_FLT_Needful    := 1,
           IN_FLT_Reset      := "DB009_Faults".Faults_Reset_FKT_M1,
           IO_Any_ArrayPV    := "DB608_PV_Metering".HeatexchangerHP[2],
           IO_Fault_Sensor   := "DB823_Error_Metering".Temperature_HeatexchangerHP[2].Sensor_FLT_broken_wire,
           IO_New_Fault      := "DB009_Faults".Faultschanging_M1,
           IO_FLT_Level_3    := "DB009_Faults".Faults_FKT_Grp_3_M1
         );
   //
         L     "DB608_PV_Metering".HeatexchangerHP[2].PV_ActV.Value;
         L     10.0;
         /R;
         T     #Temp_HD_WT;
   //
         L     "DB608_PV_Metering".HeatexchangerHP[2].PV_SetV.Value;
         L     10.0;
         /R;
         T     #Temp_SetValueTemp;
   //
         CALL  "FC056_TemPulse2"
         ( Trig              := "Start_Controler1_HP_K2",
           In_Sollwert       := #Temp_SetValueTemp,
           In_Istwert_Tank   := #Temp_HD_WT,
           In_Istwert_Return := #Temp_HD_WT,
           In_Wichtung       := "DB751_auxiliaryDriveMetering".HeatexchangerHP[2].Weighting_Temp,
           In_Regelstrecke   := "DB751_auxiliaryDriveMetering".HeatexchangerHP[2].PLC_Control_Area,
           In_MaxDelta_K     := "DB751_auxiliaryDriveMetering".HeatexchangerHP[2].Max_Temp_Diff_Cooling,
           In_MaxDelta_H     := "DB751_auxiliaryDriveMetering".HeatexchangerHP[2].Max_Temp_Diff_Heating,
           Pulsezeit         := "DB613_Komponent_State".HeatexchangerHP[2].PulsTime,
           Heating           := #Dummy,
           Cooling           := #Temp_Cooling
         );
   //
   //Regelstrecke ms Format
         L     "DB751_auxiliaryDriveMetering".HeatexchangerHP[2].PLC_Control_Area;
         L     1000.0;
         *R;
         RND;
         T     #Regelstrecke;  // Zeitwert für Timer

   // Regelstreckentimer ständig starten

         AN    "Start_Controler1_HP_K2";
         =     "Start_Controler2_HP_K2";

         CALL  TON , "DB56_Temp_HD_WT_MK1_K2"
         ( IN := "Start_Controler2_HP_K2",
           PT := #Regelstrecke,
           Q  := "Start_Controler1_HP_K2",
           ET := #Zeit_abgelaufen
         );

   // Kühlen  EIN
         A     #Temp_Cooling;
         S     "DB613_Komponent_State".HeatexchangerHP[2].CoolingActive;

   //Kleine Einschatverzögerung
         L     #Temp_SetValueTemp;
         L     "DB751_auxiliaryDriveMetering".HeatexchangerHP[2].Offset_Cooling;
         +R;
         L     #Temp_HD_WT;
         >R;
         =     #Temp_MoreDelta;

   // Kühlen  AUS
         L     "DB613_Komponent_State".HeatexchangerHP[2].PulsTime;
         RND;
         L     #Zeit_abgelaufen;
         <D;
         AN(;
         L     "DB613_Komponent_State".HeatexchangerHP[2].PulsTime;
         RND;
         L     #Regelstrecke;
         >D;
         );
         ON    "DB613_Komponent_State".HeatexchangerHP[2].Switch_Temp_ON_OFF;
         ON    "DB619_State_MPart".Operationmode[1].valid;
         O     "DB823_Error_Metering".Temperature_HeatexchangerHP[2].Sensor_FLT_broken_wire;
         O     #Temp_MoreDelta;
         R     "DB613_Komponent_State".HeatexchangerHP[2].CoolingActive;

         A     "DB613_Komponent_State".HeatexchangerHP[2].CoolingActive;
         A     "DB619_State_MPart".Machine[1].Metering."02";

         =     "V_HP_Heater_Cooling_C2";  // "V_HExchang_Cooling_K1" // stromlos zu
   //=     "V_HP_Heater_Bypass_C2" // "V_HExchang_Bypass_K1" // stromlos offen

   //-----
   // Check limits temperature 2 Heatexchanger

         CALL  "FC916_PV_Limits"
         ( IN_Tolerance_Test     := "DB619_State_MPart".Operationmode[1].Controllvoltage,
           IN_Reset_Fault        := "DB009_Faults".Faults_Reset_FKT_M1,
           IO_Any_ArrayPV        := "DB608_PV_Metering".HeatexchangerHP[2],
           IO_Fault_Warn_upperL  := "DB823_Error_Metering".Temperature_HeatexchangerHP[2].Warning_limit_plus,
           IO_Fault_Warn_lowerL  := "DB823_Error_Metering".Temperature_HeatexchangerHP[2].Warning_limit_minus,
           IO_Fault_Alarm_upperL := "DB823_Error_Metering".Temperature_HeatexchangerHP[2].Alarm_limit_plus,
           IO_Fault_Alarm_lowerL := "DB823_Error_Metering".Temperature_HeatexchangerHP[2].Alarm_limit_minus,
           IO_New_Fault          := "DB009_Faults".Faultschanging_M1,
           IO_Fault_Level_1      := "DB009_Faults".Faults_FKT_Grp_1_M1,
           IO_Fault_Level_2      := "DB009_Faults".Faults_FKT_Grp_2_M1,
           IO_Fault_Level_3      := "DB009_Faults".Faults_FKT_Grp_3_M1
         );
   //-----
   // State of Switch
         L     0;
         A     "DB613_Komponent_State".HeatexchangerHP[2].CoolingActive;
         A     "DB619_State_MPart".Machine[1].Metering."02";
         A     "DB613_Komponent_State".HeatexchangerHP[2].Switch_Temp_ON_OFF;
         JCN   S1H2;
         L     1;
   S1H2: ON    "DB613_Komponent_State".HeatexchangerHP[2].CoolingActive;
         ON    "DB619_State_MPart".Machine[1].Metering."02";
         A     "DB613_Komponent_State".HeatexchangerHP[2].Switch_Temp_ON_OFF;
         JCN   S2H2;
         L     3;
   S2H2: A     "DB823_Error_Metering".Temperature_HeatexchangerHP[2].Sensor_FLT_broken_wire;
         A     "DB613_Komponent_State".HeatexchangerHP[2].Switch_Temp_ON_OFF;
         JCN   S3H2;
         L     2;
   S3H2: T     "DB613_Komponent_State".HeatexchangerHP[2].State_Temp;
   EHD2: NOP   0;

   // Fault exists
         O     "DB823_Error_Metering".Temperature_HeatexchangerHP[2].Sensor_FLT_broken_wire;
         O     "DB823_Error_Metering".Temperature_HeatexchangerHP[2].Warning_limit_plus;
         O     "DB823_Error_Metering".Temperature_HeatexchangerHP[2].Warning_limit_minus;
         O     "DB823_Error_Metering".Temperature_HeatexchangerHP[2].Alarm_limit_plus;
         O     "DB823_Error_Metering".Temperature_HeatexchangerHP[2].Alarm_limit_minus;
         =     "DB613_Komponent_State".HeatexchangerHP[2].Fault_Exist;
END_REGION
END_FUNCTION

FUNCTION "FC057_LPHeatexchanger" : Void   // FC58, STL
{ S7_Optimized_Access := 'FALSE' }
VERSION : 0.1
   VAR_TEMP
      DINT_dummy : Real;
      Imp_WT_Aus : Bool;
      Imp_WT_Ein : Bool;
      Temp_Cooling : Bool;
      Dummy : Bool;
      Temp_MoreDelta : Bool;
      Temp_ND_WT : Real;
      Temp_SetValueTemp : Real;
      Regelstrecke : Time;
      Zeit_abgelaufen : Time;
   END_VAR
BEGIN

REGION Network 1: There is no connection to the sensor (3)
   //---------------------------------------------
   //  Controller temperature Heatexchanger K1
   //---------------------------------------------
         AN    "DB753_MeteringPump".Pump[1].WithLPHeatExchanger;
         R     "DB823_Error_Metering".Temperature_HeatexchangerLP[1].Sensor_FLT_broken_wire;
         R     "DB823_Error_Metering".Temperature_HeatexchangerLP[1].Warning_limit_plus;
         R     "DB823_Error_Metering".Temperature_HeatexchangerLP[1].Warning_limit_minus;
         R     "DB823_Error_Metering".Temperature_HeatexchangerLP[1].Alarm_limit_plus;
         R     "DB823_Error_Metering".Temperature_HeatexchangerLP[1].Alarm_limit_minus;
         R     "DB613_Komponent_State".HeatexchangerLP[1].Fault_Exist;
         JC    EHD1;
   //-----
         CALL  "FC920_PV_Calc_Act_Value"
         ( IN_Act_Value_read := TRUE,
           IN_Act_Value_ext  := FALSE,
           IN_Ext_Value      := #DINT_dummy,
           IN_Read_Double    := FALSE,
           IN_FLT_Needful    := 1,
           IN_FLT_Reset      := "DB009_Faults".Faults_Reset_FKT_M1,
           IO_Any_ArrayPV    := "DB608_PV_Metering".HeatexchangerLP[1],
           IO_Fault_Sensor   := "DB823_Error_Metering".Temperature_HeatexchangerLP[1].Sensor_FLT_broken_wire,
           IO_New_Fault      := "DB009_Faults".Faultschanging_M1,
           IO_FLT_Level_3    := "DB009_Faults".Faults_FKT_Grp_3_M1
         );

   //---------------------------------------------
   //  Controller temperature Heatexchanger K1
   //---------------------------------------------
         L     "DB608_PV_Metering".HeatexchangerLP[1].PV_ActV.Value;
         L     10.0;
         /R;
         T     #Temp_ND_WT;
   //
         L     "DB608_PV_Metering".HeatexchangerLP[1].PV_SetV.Value;
         L     10.0;
         /R;
         T     #Temp_SetValueTemp;
   //
         CALL  "FC056_TemPulse2"
         ( Trig              := "Start_Controler1_LP_K1",
           In_Sollwert       := #Temp_SetValueTemp,
           In_Istwert_Tank   := #Temp_ND_WT,
           In_Istwert_Return := #Temp_ND_WT,
           In_Wichtung       := "DB751_auxiliaryDriveMetering".HeatexchangerLP[1].Weighting_Temp,
           In_Regelstrecke   := "DB751_auxiliaryDriveMetering".HeatexchangerLP[1].PLC_Control_Area,
           In_MaxDelta_K     := "DB751_auxiliaryDriveMetering".HeatexchangerLP[1].Max_Temp_Diff_Cooling,
           In_MaxDelta_H     := "DB751_auxiliaryDriveMetering".HeatexchangerLP[1].Max_Temp_Diff_Heating,
           Pulsezeit         := "DB613_Komponent_State".HeatexchangerLP[1].PulsTime,
           Heating           := #Dummy,
           Cooling           := #Temp_Cooling
         );
   //
   //Regelstrecke ms Format
         L     "DB751_auxiliaryDriveMetering".HeatexchangerLP[1].PLC_Control_Area;
         L     1000.0;
         *R;
         RND;
         T     #Regelstrecke;  // Zeitwert für Timer

   // Regelstreckentimer ständig starten

         AN    "Start_Controler1_LP_K1";
         =     "Start_Controler2_LP_K1";

         CALL  TON , "DB60_Temp_ND_WT_MK1_K1"
         ( IN := "Start_Controler2_LP_K1",
           PT := #Regelstrecke,
           Q  := "Start_Controler1_LP_K1",
           ET := #Zeit_abgelaufen
         );

   // Kühlen  EIN
         A     #Temp_Cooling;
         S     "DB613_Komponent_State".HeatexchangerLP[1].CoolingActive;

